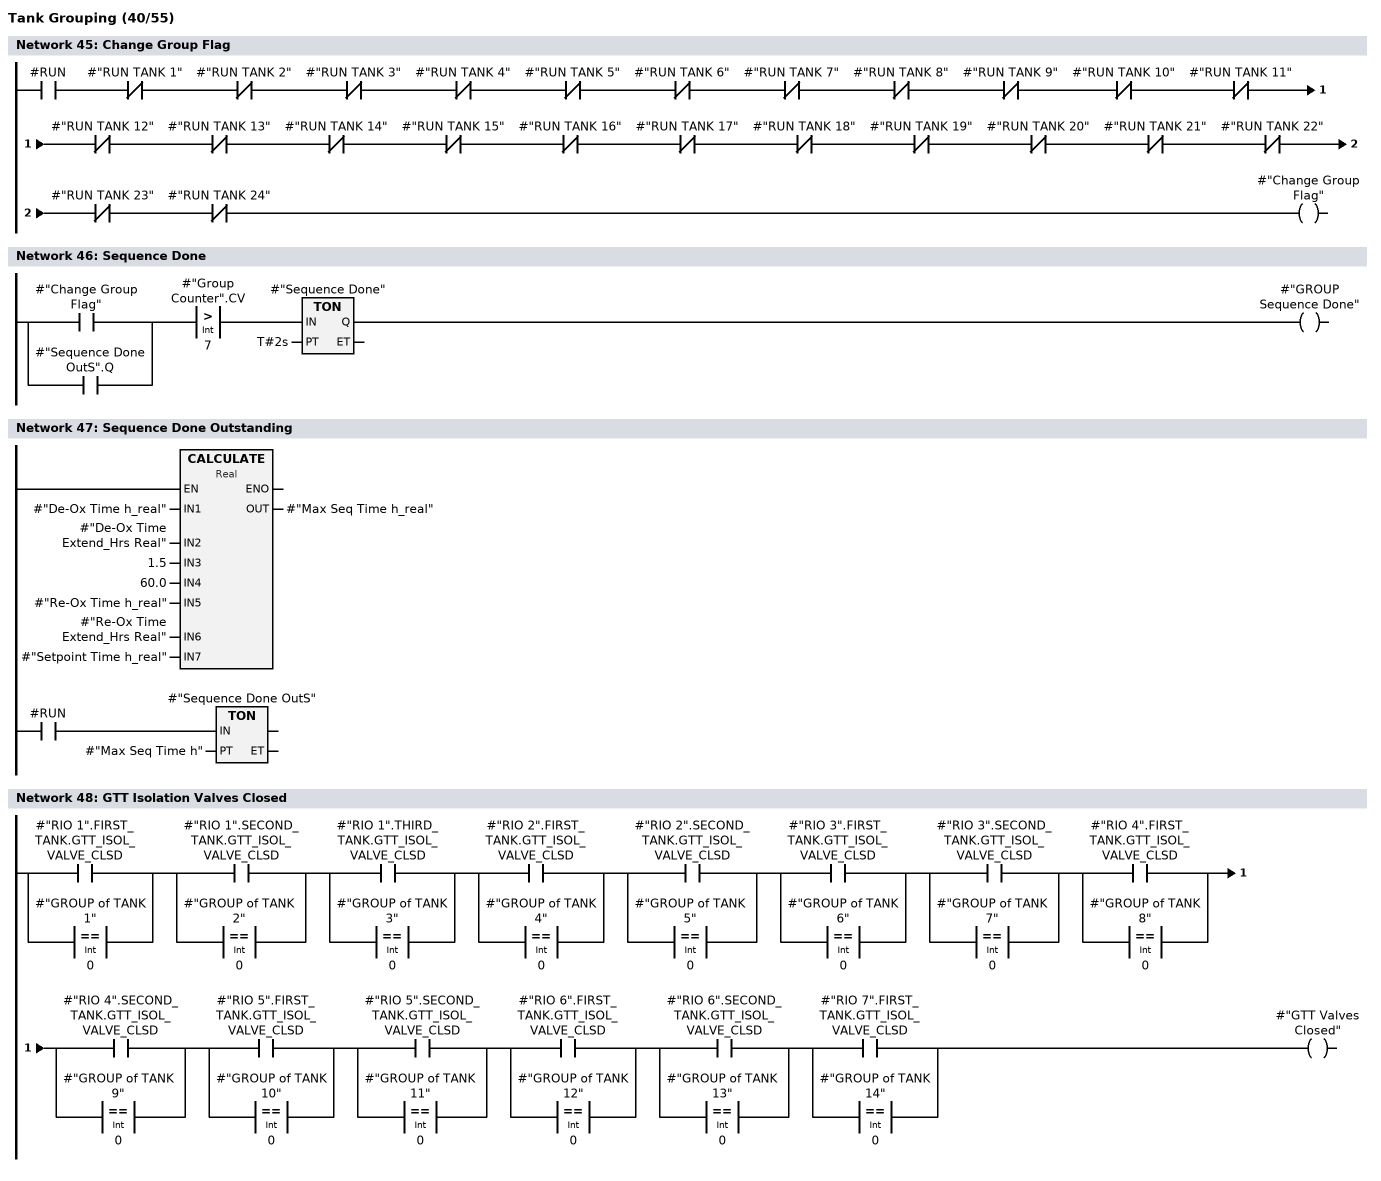
   RUNG wire#powerrail
      Contact( #RUN )
      I_Contact( #"RUN TANK 1" )
      I_Contact( #"RUN TANK 2" )
      I_Contact( #"RUN TANK 3" )
      I_Contact( #"RUN TANK 4" )
      I_Contact( #"RUN TANK 5" )
      I_Contact( #"RUN TANK 6" )
      I_Contact( #"RUN TANK 7" )
      I_Contact( #"RUN TANK 8" )
      I_Contact( #"RUN TANK 9" )
      I_Contact( #"RUN TANK 10" )
      I_Contact( #"RUN TANK 11" )
      I_Contact( #"RUN TANK 12" )
      I_Contact( #"RUN TANK 13" )
      I_Contact( #"RUN TANK 14" )
      I_Contact( #"RUN TANK 15" )
      I_Contact( #"RUN TANK 16" )
      I_Contact( #"RUN TANK 17" )
      I_Contact( #"RUN TANK 18" )
      I_Contact( #"RUN TANK 19" )
      I_Contact( #"RUN TANK 20" )
      I_Contact( #"RUN TANK 21" )
      I_Contact( #"RUN TANK 22" )
      I_Contact( #"RUN TANK 23" )
      I_Contact( #"RUN TANK 24" )
      Coil( #"Change Group Flag" )
   END_RUNG
   // the same network as SCL:
   #"Change Group Flag" := #RUN AND NOT #"RUN TANK 1" AND NOT #"RUN TANK 2" AND NOT #"RUN TANK 3" AND NOT #"RUN TANK 4" AND NOT #"RUN TANK 5" AND NOT #"RUN TANK 6" AND NOT #"RUN TANK 7" AND NOT #"RUN TANK 8" AND NOT #"RUN TANK 9" AND NOT #"RUN TANK 10" AND NOT #"RUN TANK 11" AND NOT #"RUN TANK 12" AND NOT #"RUN TANK 13" AND NOT #"RUN TANK 14" AND NOT #"RUN TANK 15" AND NOT #"RUN TANK 16" AND NOT #"RUN TANK 17" AND NOT #"RUN TANK 18" AND NOT #"RUN TANK 19" AND NOT #"RUN TANK 20" AND NOT #"RUN TANK 21" AND NOT #"RUN TANK 22" AND NOT #"RUN TANK 23" AND NOT #"RUN TANK 24";
END_REGION

REGION Network 46: Sequence Done
   #"Sequence Done"(IN := (#"Change Group Flag" OR #"Sequence Done OutS".Q) AND (#"Group Counter".CV > 7),   // TON
                    PT := T#2s);
   #"GROUP Sequence Done" := #"Sequence Done".Q;
END_REGION

REGION Network 47: Sequence Done Outstanding
   #"Max Seq Time h_real" := (#"De-Ox Time h_real"+#"De-Ox Time Extend_Hrs Real"+#"Setpoint Time h_real")*1.5;
   #"Sequence Done OutS"(IN := #RUN, PT := #"Max Seq Time h");   // TON
END_REGION

REGION Network 48: GTT Isolation Valves Closed
   RUNG wire#powerrail
      Contact( #"RIO 1".FIRST_TANK.GTT_ISOL_VALVE_CLSD )
      wire#w1
      Contact( #"RIO 1".SECOND_TANK.GTT_ISOL_VALVE_CLSD )
      wire#w2
      Contact( #"RIO 1".THIRD_TANK.GTT_ISOL_VALVE_CLSD )
      wire#w3
      Contact( #"RIO 2".FIRST_TANK.GTT_ISOL_VALVE_CLSD )
      wire#w4
      Contact( #"RIO 2".SECOND_TANK.GTT_ISOL_VALVE_CLSD )
      wire#w5
      Contact( #"RIO 3".FIRST_TANK.GTT_ISOL_VALVE_CLSD )
      wire#w6
      Contact( #"RIO 3".SECOND_TANK.GTT_ISOL_VALVE_CLSD )
      wire#w7
      Contact( #"RIO 4".FIRST_TANK.GTT_ISOL_VALVE_CLSD )
      wire#w8
      Contact( #"RIO 4".SECOND_TANK.GTT_ISOL_VALVE_CLSD )
      wire#w9
      Contact( #"RIO 5".FIRST_TANK.GTT_ISOL_VALVE_CLSD )
      wire#w10
      Contact( #"RIO 5".SECOND_TANK.GTT_ISOL_VALVE_CLSD )
      wire#w11
      Contact( #"RIO 6".FIRST_TANK.GTT_ISOL_VALVE_CLSD )
      wire#w12
      Contact( #"RIO 6".SECOND_TANK.GTT_ISOL_VALVE_CLSD )
      wire#w13
      Contact( #"RIO 7".FIRST_TANK.GTT_ISOL_VALVE_CLSD )
      wire#w14
      Coil( #"GTT Valves Closed" )
   END_RUNG
   RUNG wire#powerrail
      { S7_Templates := "SrcType := Int" } EQ_Contact(in1 := #"GROUP of TANK 1", in2 := 0)
   END_RUNG wire#w1
   RUNG wire#w1
      { S7_Templates := "SrcType := Int" } EQ_Contact(in1 := #"GROUP of TANK 2", in2 := 0)
   END_RUNG wire#w2
   RUNG wire#w2
      { S7_Templates := "SrcType := Int" } EQ_Contact(in1 := #"GROUP of TANK 3", in2 := 0)
   END_RUNG wire#w3
   RUNG wire#w3
      { S7_Templates := "SrcType := Int" } EQ_Contact(in1 := #"GROUP of TANK 4", in2 := 0)
   END_RUNG wire#w4
   RUNG wire#w4
      { S7_Templates := "SrcType := Int" } EQ_Contact(in1 := #"GROUP of TANK 5", in2 := 0)
   END_RUNG wire#w5
   RUNG wire#w5
      { S7_Templates := "SrcType := Int" } EQ_Contact(in1 := #"GROUP of TANK 6", in2 := 0)
   END_RUNG wire#w6
   RUNG wire#w6
      { S7_Templates := "SrcType := Int" } EQ_Contact(in1 := #"GROUP of TANK 7", in2 := 0)
   END_RUNG wire#w7
   RUNG wire#w7
      { S7_Templates := "SrcType := Int" } EQ_Contact(in1 := #"GROUP of TANK 8", in2 := 0)
   END_RUNG wire#w8
   RUNG wire#w8
      { S7_Templates := "SrcType := Int" } EQ_Contact(in1 := #"GROUP of TANK 9", in2 := 0)
   END_RUNG wire#w9
   RUNG wire#w9
      { S7_Templates := "SrcType := Int" } EQ_Contact(in1 := #"GROUP of TANK 10", in2 := 0)
   END_RUNG wire#w10
   RUNG wire#w10
      { S7_Templates := "SrcType := Int" } EQ_Contact(in1 := #"GROUP of TANK 11", in2 := 0)
   END_RUNG wire#w11
   RUNG wire#w11
      { S7_Templates := "SrcType := Int" } EQ_Contact(in1 := #"GROUP of TANK 12", in2 := 0)
   END_RUNG wire#w12
   RUNG wire#w12
      { S7_Templates := "SrcType := Int" } EQ_Contact(in1 := #"GROUP of TANK 13", in2 := 0)
   END_RUNG wire#w13
   RUNG wire#w13
      { S7_Templates := "SrcType := Int" } EQ_Contact(in1 := #"GROUP of TANK 14", in2 := 0)
   END_RUNG wire#w14
   // the same network as SCL:
   #"GTT Valves Closed" := (#"RIO 1".FIRST_TANK.GTT_ISOL_VALVE_CLSD OR (#"GROUP of TANK 1" = 0)) AND (#"RIO 1".SECOND_TANK.GTT_ISOL_VALVE_CLSD OR (#"GROUP of TANK 2" = 0)) AND (#"RIO 1".THIRD_TANK.GTT_ISOL_VALVE_CLSD OR (#"GROUP of TANK 3" = 0)) AND (#"RIO 2".FIRST_TANK.GTT_ISOL_VALVE_CLSD OR (#"GROUP of TANK 4" = 0)) AND (#"RIO 2".SECOND_TANK.GTT_ISOL_VALVE_CLSD OR (#"GROUP of TANK 5" = 0)) AND (#"RIO 3".FIRST_TANK.GTT_ISOL_VALVE_CLSD OR (#"GROUP of TANK 6" = 0)) AND (#"RIO 3".SECOND_TANK.GTT_ISOL_VALVE_CLSD OR (#"GROUP of TANK 7" = 0)) AND (#"RIO 4".FIRST_TANK.GTT_ISOL_VALVE_CLSD OR (#"GROUP of TANK 8" = 0)) AND (#"RIO 4".SECOND_TANK.GTT_ISOL_VALVE_CLSD OR (#"GROUP of TANK 9" = 0)) AND (#"RIO 5".FIRST_TANK.GTT_ISOL_VALVE_CLSD OR (#"GROUP of TANK 10" = 0)) AND (#"RIO 5".SECOND_TANK.GTT_ISOL_VALVE_CLSD OR (#"GROUP of TANK 11" = 0)) AND (#"RIO 6".FIRST_TANK.GTT_ISOL_VALVE_CLSD OR (#"GROUP of TANK 12" = 0)) AND (#"RIO 6".SECOND_TANK.GTT_ISOL_VALVE_CLSD OR (#"GROUP of TANK 13" = 0)) AND (#"RIO 7".FIRST_TANK.GTT_ISOL_VALVE_CLSD OR (#"GROUP of TANK 14" = 0));
END_REGION

REGION Network 49: RUN GROUP 1
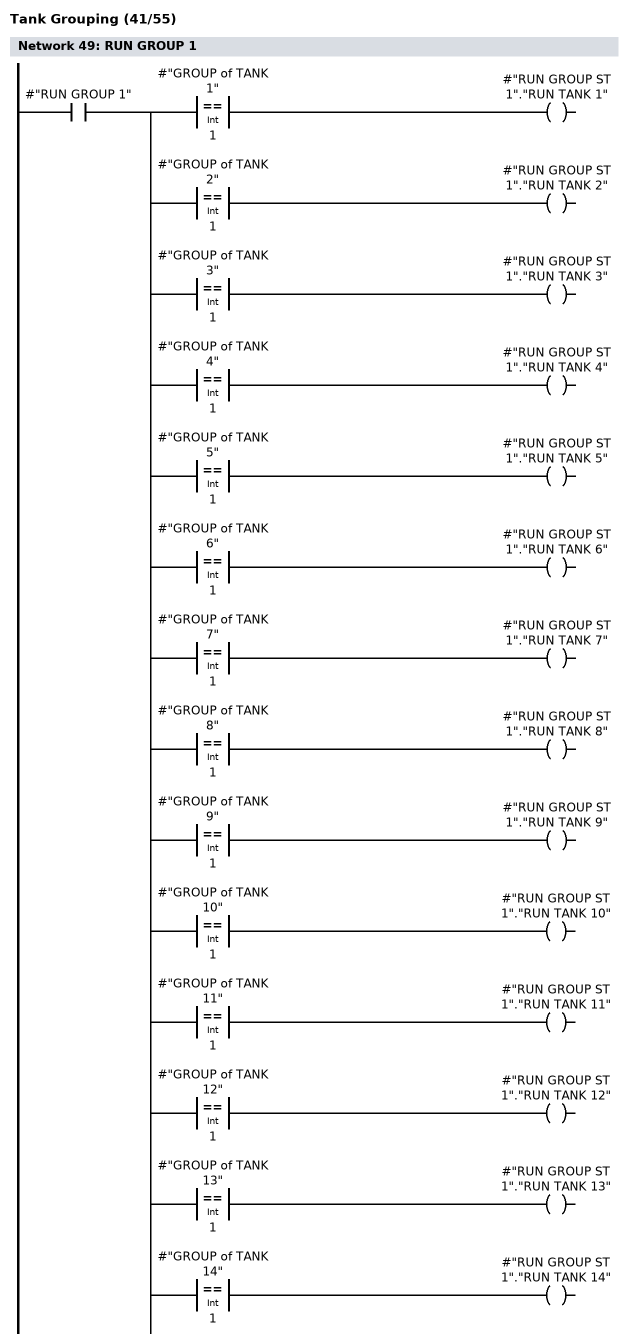
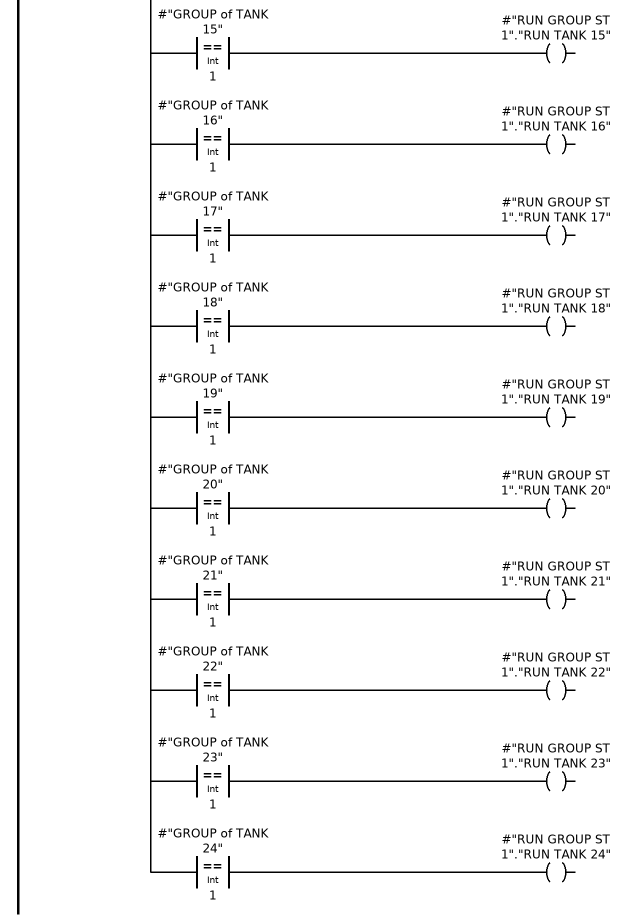
   RUNG wire#powerrail
      Contact( #"RUN GROUP 1" )
      wire#w1
      { S7_Templates := "SrcType := Int" } EQ_Contact(in1 := #"GROUP of TANK 1", in2 := 1)
      Coil( #"RUN GROUP ST 1"."RUN TANK 1" )
   END_RUNG
   RUNG wire#w1
      { S7_Templates := "SrcType := Int" } EQ_Contact(in1 := #"GROUP of TANK 2", in2 := 1)
      Coil( #"RUN GROUP ST 1"."RUN TANK 2" )
   END_RUNG
   RUNG wire#w1
      { S7_Templates := "SrcType := Int" } EQ_Contact(in1 := #"GROUP of TANK 3", in2 := 1)
      Coil( #"RUN GROUP ST 1"."RUN TANK 3" )
   END_RUNG
   RUNG wire#w1
      { S7_Templates := "SrcType := Int" } EQ_Contact(in1 := #"GROUP of TANK 4", in2 := 1)
      Coil( #"RUN GROUP ST 1"."RUN TANK 4" )
   END_RUNG
   RUNG wire#w1
      { S7_Templates := "SrcType := Int" } EQ_Contact(in1 := #"GROUP of TANK 5", in2 := 1)
      Coil( #"RUN GROUP ST 1"."RUN TANK 5" )
   END_RUNG
   RUNG wire#w1
      { S7_Templates := "SrcType := Int" } EQ_Contact(in1 := #"GROUP of TANK 6", in2 := 1)
      Coil( #"RUN GROUP ST 1"."RUN TANK 6" )
   END_RUNG
   RUNG wire#w1
      { S7_Templates := "SrcType := Int" } EQ_Contact(in1 := #"GROUP of TANK 7", in2 := 1)
      Coil( #"RUN GROUP ST 1"."RUN TANK 7" )
   END_RUNG
   RUNG wire#w1
      { S7_Templates := "SrcType := Int" } EQ_Contact(in1 := #"GROUP of TANK 8", in2 := 1)
      Coil( #"RUN GROUP ST 1"."RUN TANK 8" )
   END_RUNG
   RUNG wire#w1
      { S7_Templates := "SrcType := Int" } EQ_Contact(in1 := #"GROUP of TANK 9", in2 := 1)
      Coil( #"RUN GROUP ST 1"."RUN TANK 9" )
   END_RUNG
   RUNG wire#w1
      { S7_Templates := "SrcType := Int" } EQ_Contact(in1 := #"GROUP of TANK 10", in2 := 1)
      Coil( #"RUN GROUP ST 1"."RUN TANK 10" )
   END_RUNG
   RUNG wire#w1
      { S7_Templates := "SrcType := Int" } EQ_Contact(in1 := #"GROUP of TANK 11", in2 := 1)
      Coil( #"RUN GROUP ST 1"."RUN TANK 11" )
   END_RUNG
   RUNG wire#w1
      { S7_Templates := "SrcType := Int" } EQ_Contact(in1 := #"GROUP of TANK 12", in2 := 1)
      Coil( #"RUN GROUP ST 1"."RUN TANK 12" )
   END_RUNG
   RUNG wire#w1
      { S7_Templates := "SrcType := Int" } EQ_Contact(in1 := #"GROUP of TANK 13", in2 := 1)
      Coil( #"RUN GROUP ST 1"."RUN TANK 13" )
   END_RUNG
   RUNG wire#w1
      { S7_Templates := "SrcType := Int" } EQ_Contact(in1 := #"GROUP of TANK 14", in2 := 1)
      Coil( #"RUN GROUP ST 1"."RUN TANK 14" )
   END_RUNG
   RUNG wire#w1
      { S7_Templates := "SrcType := Int" } EQ_Contact(in1 := #"GROUP of TANK 15", in2 := 1)
      Coil( #"RUN GROUP ST 1"."RUN TANK 15" )
   END_RUNG
   RUNG wire#w1
      { S7_Templates := "SrcType := Int" } EQ_Contact(in1 := #"GROUP of TANK 16", in2 := 1)
      Coil( #"RUN GROUP ST 1"."RUN TANK 16" )
   END_RUNG
   RUNG wire#w1
      { S7_Templates := "SrcType := Int" } EQ_Contact(in1 := #"GROUP of TANK 17", in2 := 1)
      Coil( #"RUN GROUP ST 1"."RUN TANK 17" )
   END_RUNG
   RUNG wire#w1
      { S7_Templates := "SrcType := Int" } EQ_Contact(in1 := #"GROUP of TANK 18", in2 := 1)
      Coil( #"RUN GROUP ST 1"."RUN TANK 18" )
   END_RUNG
   RUNG wire#w1
      { S7_Templates := "SrcType := Int" } EQ_Contact(in1 := #"GROUP of TANK 19", in2 := 1)
      Coil( #"RUN GROUP ST 1"."RUN TANK 19" )
   END_RUNG
   RUNG wire#w1
      { S7_Templates := "SrcType := Int" } EQ_Contact(in1 := #"GROUP of TANK 20", in2 := 1)
      Coil( #"RUN GROUP ST 1"."RUN TANK 20" )
   END_RUNG
   RUNG wire#w1
      { S7_Templates := "SrcType := Int" } EQ_Contact(in1 := #"GROUP of TANK 21", in2 := 1)
      Coil( #"RUN GROUP ST 1"."RUN TANK 21" )
   END_RUNG
   RUNG wire#w1
      { S7_Templates := "SrcType := Int" } EQ_Contact(in1 := #"GROUP of TANK 22", in2 := 1)
      Coil( #"RUN GROUP ST 1"."RUN TANK 22" )
   END_RUNG
   RUNG wire#w1
      { S7_Templates := "SrcType := Int" } EQ_Contact(in1 := #"GROUP of TANK 23", in2 := 1)
      Coil( #"RUN GROUP ST 1"."RUN TANK 23" )
   END_RUNG
   RUNG wire#w1
      { S7_Templates := "SrcType := Int" } EQ_Contact(in1 := #"GROUP of TANK 24", in2 := 1)
      Coil( #"RUN GROUP ST 1"."RUN TANK 24" )
   END_RUNG
   // the same network as SCL:
   #"RUN GROUP ST 1"."RUN TANK 1" := #"RUN GROUP 1" AND (#"GROUP of TANK 1" = 1);
   #"RUN GROUP ST 1"."RUN TANK 2" := #"RUN GROUP 1" AND (#"GROUP of TANK 2" = 1);
   #"RUN GROUP ST 1"."RUN TANK 3" := #"RUN GROUP 1" AND (#"GROUP of TANK 3" = 1);
   #"RUN GROUP ST 1"."RUN TANK 4" := #"RUN GROUP 1" AND (#"GROUP of TANK 4" = 1);
   #"RUN GROUP ST 1"."RUN TANK 5" := #"RUN GROUP 1" AND (#"GROUP of TANK 5" = 1);
   #"RUN GROUP ST 1"."RUN TANK 6" := #"RUN GROUP 1" AND (#"GROUP of TANK 6" = 1);
   #"RUN GROUP ST 1"."RUN TANK 7" := #"RUN GROUP 1" AND (#"GROUP of TANK 7" = 1);
   #"RUN GROUP ST 1"."RUN TANK 8" := #"RUN GROUP 1" AND (#"GROUP of TANK 8" = 1);
   #"RUN GROUP ST 1"."RUN TANK 9" := #"RUN GROUP 1" AND (#"GROUP of TANK 9" = 1);
   #"RUN GROUP ST 1"."RUN TANK 10" := #"RUN GROUP 1" AND (#"GROUP of TANK 10" = 1);
   #"RUN GROUP ST 1"."RUN TANK 11" := #"RUN GROUP 1" AND (#"GROUP of TANK 11" = 1);
   #"RUN GROUP ST 1"."RUN TANK 12" := #"RUN GROUP 1" AND (#"GROUP of TANK 12" = 1);
   #"RUN GROUP ST 1"."RUN TANK 13" := #"RUN GROUP 1" AND (#"GROUP of TANK 13" = 1);
   #"RUN GROUP ST 1"."RUN TANK 14" := #"RUN GROUP 1" AND (#"GROUP of TANK 14" = 1);
   #"RUN GROUP ST 1"."RUN TANK 15" := #"RUN GROUP 1" AND (#"GROUP of TANK 15" = 1);
   #"RUN GROUP ST 1"."RUN TANK 16" := #"RUN GROUP 1" AND (#"GROUP of TANK 16" = 1);
   #"RUN GROUP ST 1"."RUN TANK 17" := #"RUN GROUP 1" AND (#"GROUP of TANK 17" = 1);
   #"RUN GROUP ST 1"."RUN TANK 18" := #"RUN GROUP 1" AND (#"GROUP of TANK 18" = 1);
   #"RUN GROUP ST 1"."RUN TANK 19" := #"RUN GROUP 1" AND (#"GROUP of TANK 19" = 1);
   #"RUN GROUP ST 1"."RUN TANK 20" := #"RUN GROUP 1" AND (#"GROUP of TANK 20" = 1);
   #"RUN GROUP ST 1"."RUN TANK 21" := #"RUN GROUP 1" AND (#"GROUP of TANK 21" = 1);
   #"RUN GROUP ST 1"."RUN TANK 22" := #"RUN GROUP 1" AND (#"GROUP of TANK 22" = 1);
   #"RUN GROUP ST 1"."RUN TANK 23" := #"RUN GROUP 1" AND (#"GROUP of TANK 23" = 1);
   #"RUN GROUP ST 1"."RUN TANK 24" := #"RUN GROUP 1" AND (#"GROUP of TANK 24" = 1);
END_REGION

REGION Network 50: RUN GROUP 2
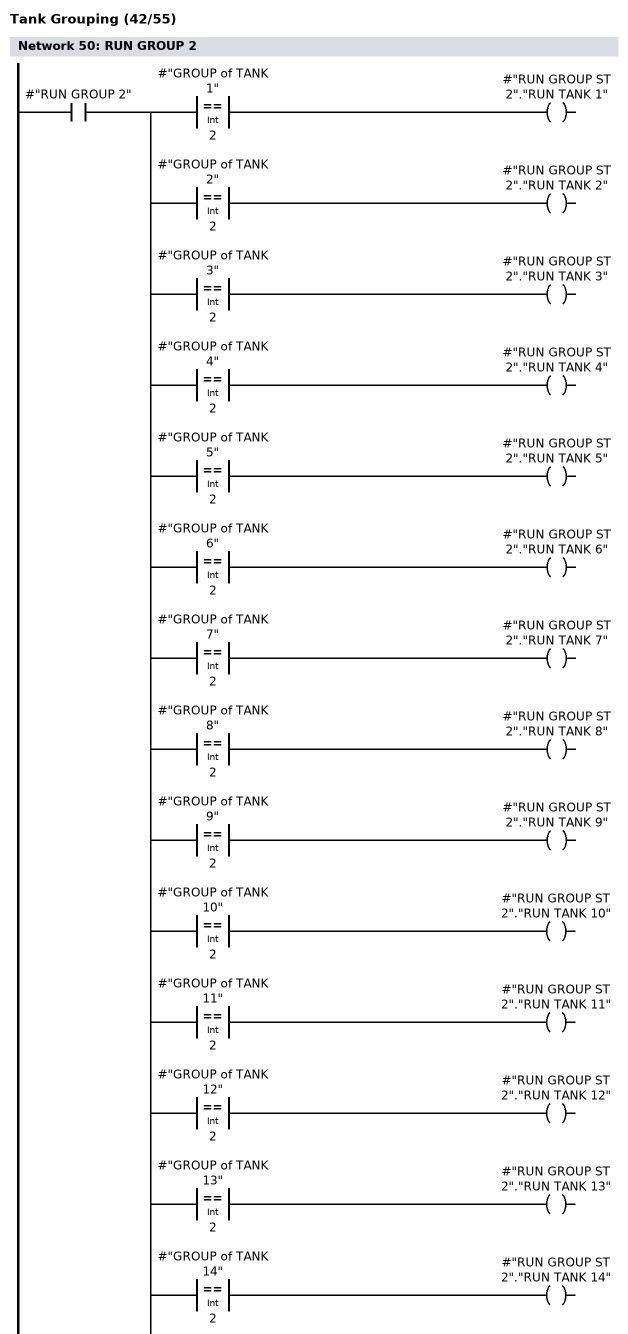
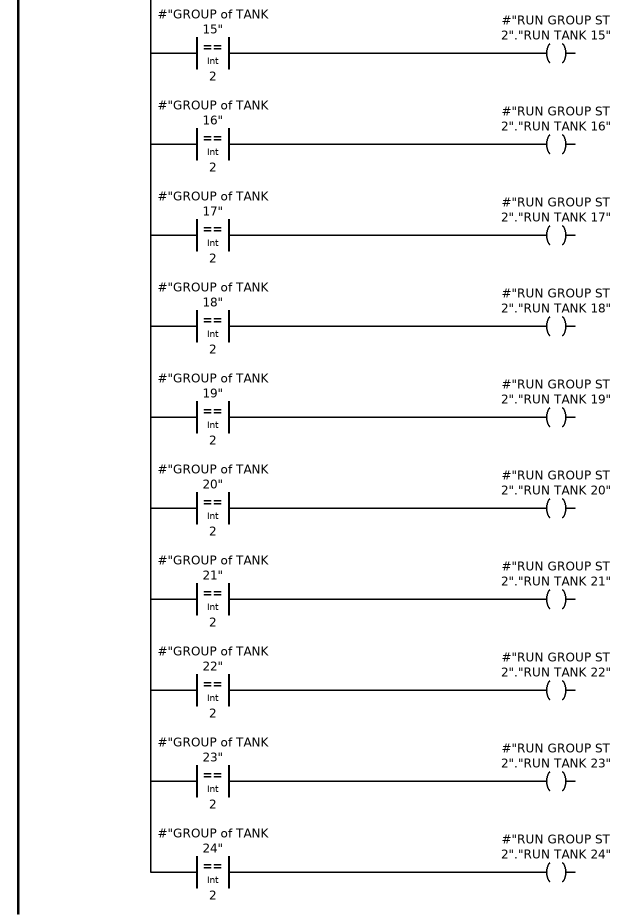
   RUNG wire#powerrail
      Contact( #"RUN GROUP 2" )
      wire#w1
      { S7_Templates := "SrcType := Int" } EQ_Contact(in1 := #"GROUP of TANK 1", in2 := 2)
      Coil( #"RUN GROUP ST 2"."RUN TANK 1" )
   END_RUNG
   RUNG wire#w1
      { S7_Templates := "SrcType := Int" } EQ_Contact(in1 := #"GROUP of TANK 2", in2 := 2)
      Coil( #"RUN GROUP ST 2"."RUN TANK 2" )
   END_RUNG
   RUNG wire#w1
      { S7_Templates := "SrcType := Int" } EQ_Contact(in1 := #"GROUP of TANK 3", in2 := 2)
      Coil( #"RUN GROUP ST 2"."RUN TANK 3" )
   END_RUNG
   RUNG wire#w1
      { S7_Templates := "SrcType := Int" } EQ_Contact(in1 := #"GROUP of TANK 4", in2 := 2)
      Coil( #"RUN GROUP ST 2"."RUN TANK 4" )
   END_RUNG
   RUNG wire#w1
      { S7_Templates := "SrcType := Int" } EQ_Contact(in1 := #"GROUP of TANK 5", in2 := 2)
      Coil( #"RUN GROUP ST 2"."RUN TANK 5" )
   END_RUNG
   RUNG wire#w1
      { S7_Templates := "SrcType := Int" } EQ_Contact(in1 := #"GROUP of TANK 6", in2 := 2)
      Coil( #"RUN GROUP ST 2"."RUN TANK 6" )
   END_RUNG
   RUNG wire#w1
      { S7_Templates := "SrcType := Int" } EQ_Contact(in1 := #"GROUP of TANK 7", in2 := 2)
      Coil( #"RUN GROUP ST 2"."RUN TANK 7" )
   END_RUNG
   RUNG wire#w1
      { S7_Templates := "SrcType := Int" } EQ_Contact(in1 := #"GROUP of TANK 8", in2 := 2)
      Coil( #"RUN GROUP ST 2"."RUN TANK 8" )
   END_RUNG
   RUNG wire#w1
      { S7_Templates := "SrcType := Int" } EQ_Contact(in1 := #"GROUP of TANK 9", in2 := 2)
      Coil( #"RUN GROUP ST 2"."RUN TANK 9" )
   END_RUNG
   RUNG wire#w1
      { S7_Templates := "SrcType := Int" } EQ_Contact(in1 := #"GROUP of TANK 10", in2 := 2)
      Coil( #"RUN GROUP ST 2"."RUN TANK 10" )
   END_RUNG
   RUNG wire#w1
      { S7_Templates := "SrcType := Int" } EQ_Contact(in1 := #"GROUP of TANK 11", in2 := 2)
      Coil( #"RUN GROUP ST 2"."RUN TANK 11" )
   END_RUNG
   RUNG wire#w1
      { S7_Templates := "SrcType := Int" } EQ_Contact(in1 := #"GROUP of TANK 12", in2 := 2)
      Coil( #"RUN GROUP ST 2"."RUN TANK 12" )
   END_RUNG
   RUNG wire#w1
      { S7_Templates := "SrcType := Int" } EQ_Contact(in1 := #"GROUP of TANK 13", in2 := 2)
      Coil( #"RUN GROUP ST 2"."RUN TANK 13" )
   END_RUNG
   RUNG wire#w1
      { S7_Templates := "SrcType := Int" } EQ_Contact(in1 := #"GROUP of TANK 14", in2 := 2)
      Coil( #"RUN GROUP ST 2"."RUN TANK 14" )
   END_RUNG
   RUNG wire#w1
      { S7_Templates := "SrcType := Int" } EQ_Contact(in1 := #"GROUP of TANK 15", in2 := 2)
      Coil( #"RUN GROUP ST 2"."RUN TANK 15" )
   END_RUNG
   RUNG wire#w1
      { S7_Templates := "SrcType := Int" } EQ_Contact(in1 := #"GROUP of TANK 16", in2 := 2)
      Coil( #"RUN GROUP ST 2"."RUN TANK 16" )
   END_RUNG
   RUNG wire#w1
      { S7_Templates := "SrcType := Int" } EQ_Contact(in1 := #"GROUP of TANK 17", in2 := 2)
      Coil( #"RUN GROUP ST 2"."RUN TANK 17" )
   END_RUNG
   RUNG wire#w1
      { S7_Templates := "SrcType := Int" } EQ_Contact(in1 := #"GROUP of TANK 18", in2 := 2)
      Coil( #"RUN GROUP ST 2"."RUN TANK 18" )
   END_RUNG
   RUNG wire#w1
      { S7_Templates := "SrcType := Int" } EQ_Contact(in1 := #"GROUP of TANK 19", in2 := 2)
      Coil( #"RUN GROUP ST 2"."RUN TANK 19" )
   END_RUNG
   RUNG wire#w1
      { S7_Templates := "SrcType := Int" } EQ_Contact(in1 := #"GROUP of TANK 20", in2 := 2)
      Coil( #"RUN GROUP ST 2"."RUN TANK 20" )
   END_RUNG
   RUNG wire#w1
      { S7_Templates := "SrcType := Int" } EQ_Contact(in1 := #"GROUP of TANK 21", in2 := 2)
      Coil( #"RUN GROUP ST 2"."RUN TANK 21" )
   END_RUNG
   RUNG wire#w1
      { S7_Templates := "SrcType := Int" } EQ_Contact(in1 := #"GROUP of TANK 22", in2 := 2)
      Coil( #"RUN GROUP ST 2"."RUN TANK 22" )
   END_RUNG
   RUNG wire#w1
      { S7_Templates := "SrcType := Int" } EQ_Contact(in1 := #"GROUP of TANK 23", in2 := 2)
      Coil( #"RUN GROUP ST 2"."RUN TANK 23" )
   END_RUNG
   RUNG wire#w1
      { S7_Templates := "SrcType := Int" } EQ_Contact(in1 := #"GROUP of TANK 24", in2 := 2)
      Coil( #"RUN GROUP ST 2"."RUN TANK 24" )
   END_RUNG
   // the same network as SCL:
   #"RUN GROUP ST 2"."RUN TANK 1" := #"RUN GROUP 2" AND (#"GROUP of TANK 1" = 2);
   #"RUN GROUP ST 2"."RUN TANK 2" := #"RUN GROUP 2" AND (#"GROUP of TANK 2" = 2);
   #"RUN GROUP ST 2"."RUN TANK 3" := #"RUN GROUP 2" AND (#"GROUP of TANK 3" = 2);
   #"RUN GROUP ST 2"."RUN TANK 4" := #"RUN GROUP 2" AND (#"GROUP of TANK 4" = 2);
   #"RUN GROUP ST 2"."RUN TANK 5" := #"RUN GROUP 2" AND (#"GROUP of TANK 5" = 2);
   #"RUN GROUP ST 2"."RUN TANK 6" := #"RUN GROUP 2" AND (#"GROUP of TANK 6" = 2);
   #"RUN GROUP ST 2"."RUN TANK 7" := #"RUN GROUP 2" AND (#"GROUP of TANK 7" = 2);
   #"RUN GROUP ST 2"."RUN TANK 8" := #"RUN GROUP 2" AND (#"GROUP of TANK 8" = 2);
   #"RUN GROUP ST 2"."RUN TANK 9" := #"RUN GROUP 2" AND (#"GROUP of TANK 9" = 2);
   #"RUN GROUP ST 2"."RUN TANK 10" := #"RUN GROUP 2" AND (#"GROUP of TANK 10" = 2);
   #"RUN GROUP ST 2"."RUN TANK 11" := #"RUN GROUP 2" AND (#"GROUP of TANK 11" = 2);
   #"RUN GROUP ST 2"."RUN TANK 12" := #"RUN GROUP 2" AND (#"GROUP of TANK 12" = 2);
   #"RUN GROUP ST 2"."RUN TANK 13" := #"RUN GROUP 2" AND (#"GROUP of TANK 13" = 2);
   #"RUN GROUP ST 2"."RUN TANK 14" := #"RUN GROUP 2" AND (#"GROUP of TANK 14" = 2);
   #"RUN GROUP ST 2"."RUN TANK 15" := #"RUN GROUP 2" AND (#"GROUP of TANK 15" = 2);
   #"RUN GROUP ST 2"."RUN TANK 16" := #"RUN GROUP 2" AND (#"GROUP of TANK 16" = 2);
   #"RUN GROUP ST 2"."RUN TANK 17" := #"RUN GROUP 2" AND (#"GROUP of TANK 17" = 2);
   #"RUN GROUP ST 2"."RUN TANK 18" := #"RUN GROUP 2" AND (#"GROUP of TANK 18" = 2);
   #"RUN GROUP ST 2"."RUN TANK 19" := #"RUN GROUP 2" AND (#"GROUP of TANK 19" = 2);
   #"RUN GROUP ST 2"."RUN TANK 20" := #"RUN GROUP 2" AND (#"GROUP of TANK 20" = 2);
   #"RUN GROUP ST 2"."RUN TANK 21" := #"RUN GROUP 2" AND (#"GROUP of TANK 21" = 2);
   #"RUN GROUP ST 2"."RUN TANK 22" := #"RUN GROUP 2" AND (#"GROUP of TANK 22" = 2);
   #"RUN GROUP ST 2"."RUN TANK 23" := #"RUN GROUP 2" AND (#"GROUP of TANK 23" = 2);
   #"RUN GROUP ST 2"."RUN TANK 24" := #"RUN GROUP 2" AND (#"GROUP of TANK 24" = 2);
END_REGION

REGION Network 51: RUN GROUP 3
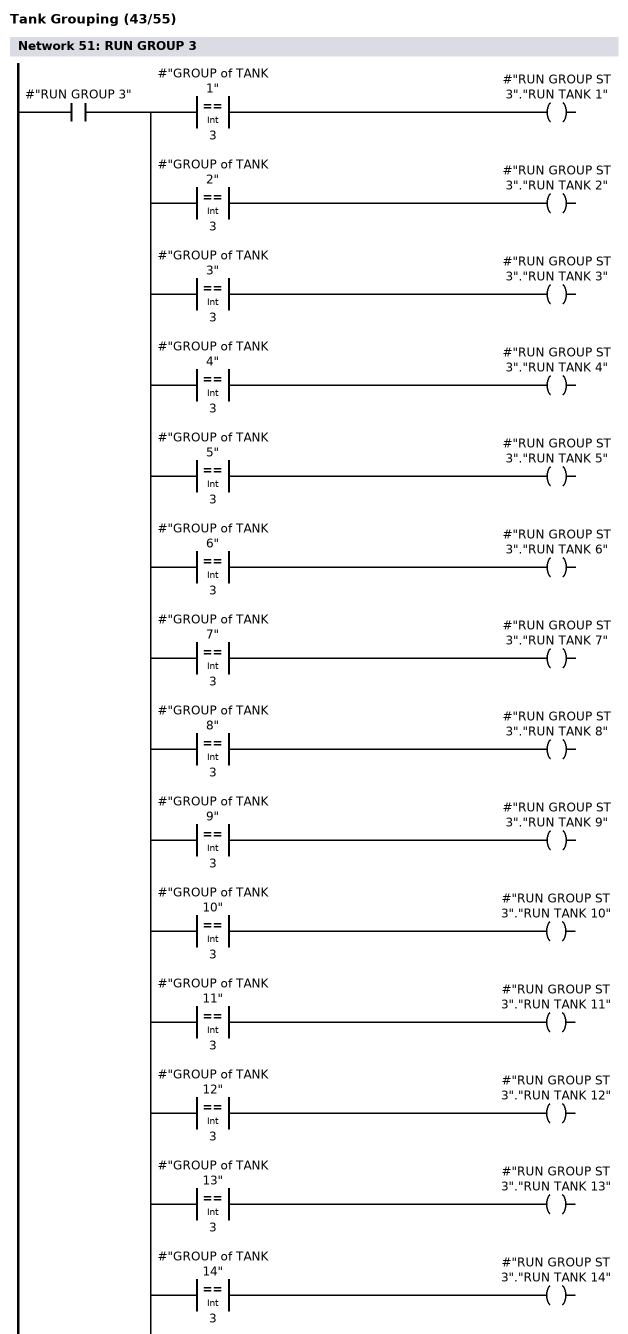
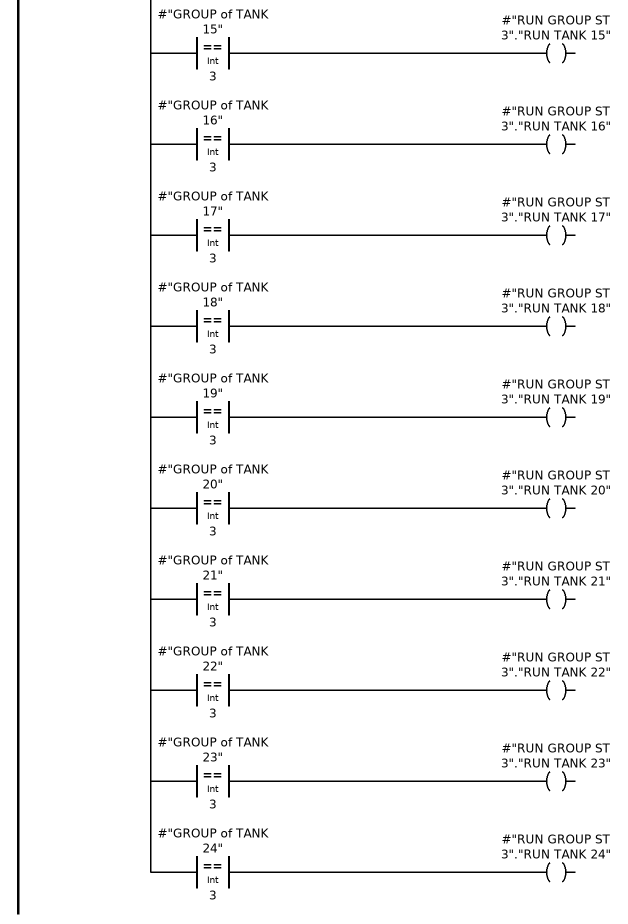
   RUNG wire#powerrail
      Contact( #"RUN GROUP 3" )
      wire#w1
      { S7_Templates := "SrcType := Int" } EQ_Contact(in1 := #"GROUP of TANK 1", in2 := 3)
      Coil( #"RUN GROUP ST 3"."RUN TANK 1" )
   END_RUNG
   RUNG wire#w1
      { S7_Templates := "SrcType := Int" } EQ_Contact(in1 := #"GROUP of TANK 2", in2 := 3)
      Coil( #"RUN GROUP ST 3"."RUN TANK 2" )
   END_RUNG
   RUNG wire#w1
      { S7_Templates := "SrcType := Int" } EQ_Contact(in1 := #"GROUP of TANK 3", in2 := 3)
      Coil( #"RUN GROUP ST 3"."RUN TANK 3" )
   END_RUNG
   RUNG wire#w1
      { S7_Templates := "SrcType := Int" } EQ_Contact(in1 := #"GROUP of TANK 4", in2 := 3)
      Coil( #"RUN GROUP ST 3"."RUN TANK 4" )
   END_RUNG
   RUNG wire#w1
      { S7_Templates := "SrcType := Int" } EQ_Contact(in1 := #"GROUP of TANK 5", in2 := 3)
      Coil( #"RUN GROUP ST 3"."RUN TANK 5" )
   END_RUNG
   RUNG wire#w1
      { S7_Templates := "SrcType := Int" } EQ_Contact(in1 := #"GROUP of TANK 6", in2 := 3)
      Coil( #"RUN GROUP ST 3"."RUN TANK 6" )
   END_RUNG
   RUNG wire#w1
      { S7_Templates := "SrcType := Int" } EQ_Contact(in1 := #"GROUP of TANK 7", in2 := 3)
      Coil( #"RUN GROUP ST 3"."RUN TANK 7" )
   END_RUNG
   RUNG wire#w1
      { S7_Templates := "SrcType := Int" } EQ_Contact(in1 := #"GROUP of TANK 8", in2 := 3)
      Coil( #"RUN GROUP ST 3"."RUN TANK 8" )
   END_RUNG
   RUNG wire#w1
      { S7_Templates := "SrcType := Int" } EQ_Contact(in1 := #"GROUP of TANK 9", in2 := 3)
      Coil( #"RUN GROUP ST 3"."RUN TANK 9" )
   END_RUNG
   RUNG wire#w1
      { S7_Templates := "SrcType := Int" } EQ_Contact(in1 := #"GROUP of TANK 10", in2 := 3)
      Coil( #"RUN GROUP ST 3"."RUN TANK 10" )
   END_RUNG
   RUNG wire#w1
      { S7_Templates := "SrcType := Int" } EQ_Contact(in1 := #"GROUP of TANK 11", in2 := 3)
      Coil( #"RUN GROUP ST 3"."RUN TANK 11" )
   END_RUNG
   RUNG wire#w1
      { S7_Templates := "SrcType := Int" } EQ_Contact(in1 := #"GROUP of TANK 12", in2 := 3)
      Coil( #"RUN GROUP ST 3"."RUN TANK 12" )
   END_RUNG
   RUNG wire#w1
      { S7_Templates := "SrcType := Int" } EQ_Contact(in1 := #"GROUP of TANK 13", in2 := 3)
      Coil( #"RUN GROUP ST 3"."RUN TANK 13" )
   END_RUNG
   RUNG wire#w1
      { S7_Templates := "SrcType := Int" } EQ_Contact(in1 := #"GROUP of TANK 14", in2 := 3)
      Coil( #"RUN GROUP ST 3"."RUN TANK 14" )
   END_RUNG
   RUNG wire#w1
      { S7_Templates := "SrcType := Int" } EQ_Contact(in1 := #"GROUP of TANK 15", in2 := 3)
      Coil( #"RUN GROUP ST 3"."RUN TANK 15" )
   END_RUNG
   RUNG wire#w1
      { S7_Templates := "SrcType := Int" } EQ_Contact(in1 := #"GROUP of TANK 16", in2 := 3)
      Coil( #"RUN GROUP ST 3"."RUN TANK 16" )
   END_RUNG
   RUNG wire#w1
      { S7_Templates := "SrcType := Int" } EQ_Contact(in1 := #"GROUP of TANK 17", in2 := 3)
      Coil( #"RUN GROUP ST 3"."RUN TANK 17" )
   END_RUNG
   RUNG wire#w1
      { S7_Templates := "SrcType := Int" } EQ_Contact(in1 := #"GROUP of TANK 18", in2 := 3)
      Coil( #"RUN GROUP ST 3"."RUN TANK 18" )
   END_RUNG
   RUNG wire#w1
      { S7_Templates := "SrcType := Int" } EQ_Contact(in1 := #"GROUP of TANK 19", in2 := 3)
      Coil( #"RUN GROUP ST 3"."RUN TANK 19" )
   END_RUNG
   RUNG wire#w1
      { S7_Templates := "SrcType := Int" } EQ_Contact(in1 := #"GROUP of TANK 20", in2 := 3)
      Coil( #"RUN GROUP ST 3"."RUN TANK 20" )
   END_RUNG
   RUNG wire#w1
      { S7_Templates := "SrcType := Int" } EQ_Contact(in1 := #"GROUP of TANK 21", in2 := 3)
      Coil( #"RUN GROUP ST 3"."RUN TANK 21" )
   END_RUNG
   RUNG wire#w1
      { S7_Templates := "SrcType := Int" } EQ_Contact(in1 := #"GROUP of TANK 22", in2 := 3)
      Coil( #"RUN GROUP ST 3"."RUN TANK 22" )
   END_RUNG
   RUNG wire#w1
      { S7_Templates := "SrcType := Int" } EQ_Contact(in1 := #"GROUP of TANK 23", in2 := 3)
      Coil( #"RUN GROUP ST 3"."RUN TANK 23" )
   END_RUNG
   RUNG wire#w1
      { S7_Templates := "SrcType := Int" } EQ_Contact(in1 := #"GROUP of TANK 24", in2 := 3)
      Coil( #"RUN GROUP ST 3"."RUN TANK 24" )
   END_RUNG
   // the same network as SCL:
   #"RUN GROUP ST 3"."RUN TANK 1" := #"RUN GROUP 3" AND (#"GROUP of TANK 1" = 3);
   #"RUN GROUP ST 3"."RUN TANK 2" := #"RUN GROUP 3" AND (#"GROUP of TANK 2" = 3);
   #"RUN GROUP ST 3"."RUN TANK 3" := #"RUN GROUP 3" AND (#"GROUP of TANK 3" = 3);
   #"RUN GROUP ST 3"."RUN TANK 4" := #"RUN GROUP 3" AND (#"GROUP of TANK 4" = 3);
   #"RUN GROUP ST 3"."RUN TANK 5" := #"RUN GROUP 3" AND (#"GROUP of TANK 5" = 3);
   #"RUN GROUP ST 3"."RUN TANK 6" := #"RUN GROUP 3" AND (#"GROUP of TANK 6" = 3);
   #"RUN GROUP ST 3"."RUN TANK 7" := #"RUN GROUP 3" AND (#"GROUP of TANK 7" = 3);
   #"RUN GROUP ST 3"."RUN TANK 8" := #"RUN GROUP 3" AND (#"GROUP of TANK 8" = 3);
   #"RUN GROUP ST 3"."RUN TANK 9" := #"RUN GROUP 3" AND (#"GROUP of TANK 9" = 3);
   #"RUN GROUP ST 3"."RUN TANK 10" := #"RUN GROUP 3" AND (#"GROUP of TANK 10" = 3);
   #"RUN GROUP ST 3"."RUN TANK 11" := #"RUN GROUP 3" AND (#"GROUP of TANK 11" = 3);
   #"RUN GROUP ST 3"."RUN TANK 12" := #"RUN GROUP 3" AND (#"GROUP of TANK 12" = 3);
   #"RUN GROUP ST 3"."RUN TANK 13" := #"RUN GROUP 3" AND (#"GROUP of TANK 13" = 3);
   #"RUN GROUP ST 3"."RUN TANK 14" := #"RUN GROUP 3" AND (#"GROUP of TANK 14" = 3);
   #"RUN GROUP ST 3"."RUN TANK 15" := #"RUN GROUP 3" AND (#"GROUP of TANK 15" = 3);
   #"RUN GROUP ST 3"."RUN TANK 16" := #"RUN GROUP 3" AND (#"GROUP of TANK 16" = 3);
   #"RUN GROUP ST 3"."RUN TANK 17" := #"RUN GROUP 3" AND (#"GROUP of TANK 17" = 3);
   #"RUN GROUP ST 3"."RUN TANK 18" := #"RUN GROUP 3" AND (#"GROUP of TANK 18" = 3);
   #"RUN GROUP ST 3"."RUN TANK 19" := #"RUN GROUP 3" AND (#"GROUP of TANK 19" = 3);
   #"RUN GROUP ST 3"."RUN TANK 20" := #"RUN GROUP 3" AND (#"GROUP of TANK 20" = 3);
   #"RUN GROUP ST 3"."RUN TANK 21" := #"RUN GROUP 3" AND (#"GROUP of TANK 21" = 3);
   #"RUN GROUP ST 3"."RUN TANK 22" := #"RUN GROUP 3" AND (#"GROUP of TANK 22" = 3);
   #"RUN GROUP ST 3"."RUN TANK 23" := #"RUN GROUP 3" AND (#"GROUP of TANK 23" = 3);
   #"RUN GROUP ST 3"."RUN TANK 24" := #"RUN GROUP 3" AND (#"GROUP of TANK 24" = 3);
END_REGION

REGION Network 52: RUN GROUP 4
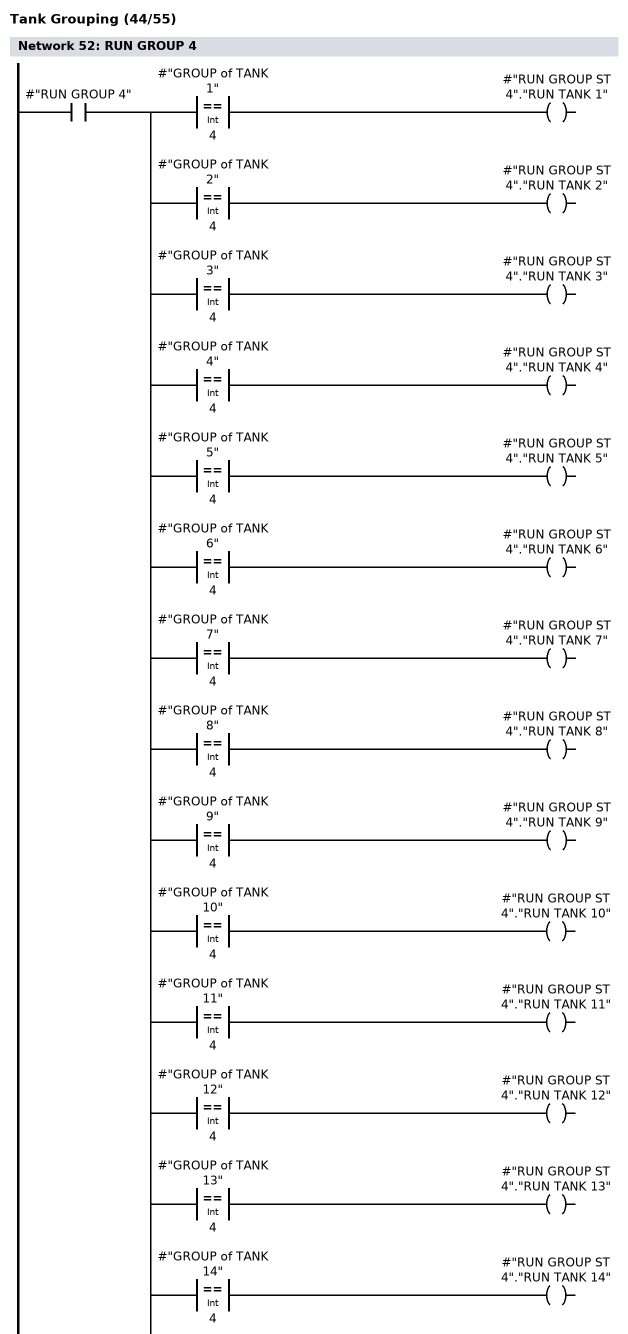
